TYPE "UDT_Segment"
VERSION : 0.1
   STRUCT
      MC_No_new : Byte := B#16#0;
      MC_No_old : Byte := B#16#0;
      Adresse_Peripherie : Word := W#16#0;
      Stationnumber : Byte := B#16#0;
      Spare_Byte_005 : Byte := B#16#0;
      Adr_Peripherie_analog : Word := W#16#0;
      Adr_Peripherie_SiemensFC : Word := W#16#0;
      Segment : "UDT_Station";
      Spare_Word_014 : Word := W#16#0;
      Spare_Word_016 : Word := W#16#0;
      Spare_Word_018 : Word := W#16#0;
      Input_from_segment : "UDT_Seg_input";
      Output_to_segment : "UDT_Seg_output";
      Siemens : "UDT_Siemens";
      Spare_Word_028 : Word := W#16#0;
      Spare_Word_030 : Word := W#16#0;
      Spare_Word_032 : Word := W#16#0;
      Spare_Word_034 : Word := W#16#0;
      Spare_Word_036 : Word := W#16#0;
      Spare_Word_038 : Word := W#16#0;
      Analogvalue_tool : Struct
         Input_lower_tool_1 : Word;
         Input_lower_tool_2 : Word;
         Input_upper_tool_1 : Word;
         Input_upper_tool_2 : Word;
      END_STRUCT;
      Input_from_tool : "UDT_Tool_Inputs_type_1";
      Output_to_tool : "UDT_Tool_Outputs_type_1";
      State_tool : "UDT_Mould_status";
      Spare_Word_068 : Word := W#16#0;
      Spare_Word_070 : Word := W#16#0;
      Spare_Word_072 : Word := W#16#0;
      Spare_Word_074 : Word := W#16#0;
      Spare_Word_076 : Word := W#16#0;
      Spare_Word_078 : Word := W#16#0;
      Spare_Word_080 : Word := W#16#0;
      Spare_Word_082 : Word := W#16#0;
      Spare_Word_084 : Word := W#16#0;
      Spare_Word_086 : Word := W#16#0;
      Spare_Word_088 : Word := W#16#0;
      Spare_Word_090 : Word := W#16#0;
      Spare_Word_092 : Word := W#16#0;
      Spare_Word_094 : Word := W#16#0;
      Spare_Word_096 : Word := W#16#0;
      Spare_Word_098 : Word := W#16#0;
      Segment_Bits : Struct
         WW_angewaehlt : Bool;
         Teachen_angewaehlt : Bool;
         STG_Nummer_wechselt : Bool;
         Nummer_geloescht : Bool;
         Beflammen_angewaehlt : Bool;
         Flag_TT_not_in_position : Bool;
         Reserve_100_6 : Bool;
         Reserve_100_7 : Bool;
         Reserve_101_0 : Bool;
         Reserve_101_1 : Bool;
         Reserve_101_2 : Bool;
         Reserve_101_3 : Bool;
         Reserve_101_4 : Bool;
         Reserve_101_5 : Bool;
         Reserve_101_6 : Bool;
         Reserve_101_7 : Bool;
         Reserve_Word_102 : Word;
         Reserve_Word_104 : Word;
         Reserve_Word_106 : Word;
         Reserve_Word_108 : Word;
      END_STRUCT;
      State_MC : Struct
         Movement : Struct
            RequestFromOP : "UDT_Actions";
            Request : "UDT_Actions";
            Command : "UDT_Actions";
            Valve : "UDT_Actions";
            End : "UDT_Actions";
         END_STRUCT;
         Cycle : "UDT_Cycle";
         Vacuum : "UDT_Vacuum";
         Seals : Struct
            Request_seal : Struct
               "1" : Bool;
               "2" : Bool;
               "3" : Bool;
               "4" : Bool;
               "5" : Bool;
               "6" : Bool;
               "7" : Bool;
               "8" : Bool;
               "9" : Bool;
               "10" : Bool;
               "11" : Bool;
               "12" : Bool;
               "13" : Bool;
               "14" : Bool;
               "15" : Bool;
               "16" : Bool;
               "17" : Bool;
               "18" : Bool;
               "19" : Bool;
               "20" : Bool;
               "21" : Bool;
               "22" : Bool;
               "23" : Bool;
               "24" : Bool;
               "25" : Bool;
               "26" : Bool;
               "27" : Bool;
               "28" : Bool;
               "29" : Bool;
               "30" : Bool;
               "31" : Bool;
               "32" : Bool;
            END_STRUCT;
            Seal_active : Array[0..32] of Byte;
            Flow : Struct
               Act_flow_1 : Real;
               Act_flow_2 : Real;
               Act_flow_3 : Real;
               Seal_faulty : Bool;
               Spare_12_1 : Bool;
               Spare_12_2 : Bool;
               Spare_12_3 : Bool;
               Spare_12_4 : Bool;
               Spare_12_5 : Bool;
               Spare_12_6 : Bool;
               Spare_12_7 : Bool;
               Spare_13_0 : Bool;
               Spare_13_1 : Bool;
               Spare_13_2 : Bool;
               Spare_13_3 : Bool;
               Spare_13_4 : Bool;
               Spare_13_5 : Bool;
               Spare_13_6 : Bool;
               Spare_13_7 : Bool;
            END_STRUCT;
         END_STRUCT;
         Operating_panel : Struct
            State : Struct
               Hydraulic_running : Bool := false;
               without_lockings : Bool := false;
               Spare_0_2 : Bool;
               Spare_0_3 : Bool;
               Spare_0_4 : Bool;
               Spare_0_5 : Bool;
               Spare_0_6 : Bool;
               Spare_0_7 : Bool;
               Act_step_program : Int := 0;   // Running, interupted or, for tool change: finished, running
               State_act_program : Int := 0;
               Act_operating_hours : Int := 0;
               Movement_blocked : Int := 0;
               Movement_condition_missing : Int := 0;
               Code_tool_01_actual : Int := 0;
               Code_tool_02_actual : Int := 0;
               Act_program : Int := 0;
               CounterMCCycles : DInt := L#1;
               DayCounterMCCycles : DInt := L#1;
               Act_cycle_time : Int := 0;
               Last_cycle_time : Int;
               Data_actual_MC : Int := 1;
               ProgStepNo : Int := 0;
               ProgType : Int := 5;
               Start_VNC : Bool := false;   // Bit to start the VNC viewer from PLC
               Fault_groupe_1_active : Bool := false;
               Fault_groupe_2_active : Bool := false;
               Fault_groupe_3_active : Bool := false;
               Fault_groupe_4_active : Bool := false;
               Check_USB : Bool := false;
               Spare_38_6 : Bool;
               Spare_38_7 : Bool;
            END_STRUCT;
            Set : Struct
               Insert_prog_line : Bool := false;
               Delete_prog_line : Bool := false;
               Movement_requested : Bool := false;
               Spare_0_3 : Bool := false;
               Spare_0_4 : Bool := false;
               Spare_0_5 : Bool := false;
               Request_search_missing_mov_cond : Bool := false;
               Search_missing_mov_cond : Bool := false;
               Start_loading_files : Bool := false;   // Starting loading files TP
               Loading_finished_TP : Bool := false;   // Loading finished TP (script finish)
               Loading_finished_PLC : Bool := false;   // Loading finished PLC (data in the plc)
               Request_write : Bool := false;   // Request signal to plc to write the next data block
               Release_write : Bool := false;   // Release signal to HMI (Script) to write the next data block
               Spare_1_5 : Bool := false;
               Spare_1_6 : Bool := false;
               Quit_fault : Bool := false;
               Selected_datablock : Int := 17;
               Selected_prog_line : Int := 49;
               Data_select : Int := 0;
               Data_actual : Int := 0;
               Selected_Axis : Int;
               User_level : Int;   // User level from HMI
               Spare_48_0 : Bool;
               Jog_axis_slow : Bool;   // Slow jog mode for referencing
               Jog_axis : Bool := false;
               Simmulate_tool : Bool := false;   // Simulate a tool. Reset in OB100! Only for testing
               Toggle_Lebensbit : Bool := false;
               Test_run_IBN : Bool;   // Test run for commisioning
               Spare_10_6 : Bool;
               Spare_10_7 : Bool;
               Act_file_name : String[30];
            END_STRUCT;
         END_STRUCT;
         Act_times : Struct
            Reaction_time_1 : Time;
            Reaction_time_2 : Time := T#0ms;
            Reaction_time_3 : Time := T#0ms;
            Reaction_time_4 : Time := T#0ms;
            Reaction_time_5 : Time := T#0ms;
            Reaction_time_6 : Time := T#0ms;
            Time_befor_degasing_tool_1 : Time := T#0ms;
            Degasing_time_tool_1 : Time := T#0ms;
            Time_befor_degasing_tool_2 : Time := T#0ms;
            Degasing_time_tool_2 : Time := T#0ms;
            Time_befor_degasing_tool_3 : Time := T#0ms;
            Degasing_time_tool_3 : Time := T#0ms;
            Time_befor_degasing_tool_4 : Time := T#0ms;
            Degasing_time_tool_4 : Time := T#0ms;
            Time_befor_degasing_tool_5 : Time := T#0ms;
            Degasing_time_tool_5 : Time := T#0ms;
            Time_befor_degasing_tool_6 : Time := T#0ms;
            Degasing_time_tool_6 : Time := T#0ms;
            Waiting_time_1 : Time := T#0ms;
            Waiting_time_2 : Time := T#0ms;
            Waiting_time_3 : Time := T#0ms;
            Waiting_time_4 : Time := T#0ms;
            Waiting_time_5 : Time := T#0ms;
            Waiting_time_6 : Time := T#0ms;
            Test_vacuum_circit_1 : Time := T#0ms;   // Dauer des Vakuumtestes für den Vakuumkreis 01
            Test_vacuum_circit_2 : Time := T#0ms;   // Dauer des Vakuumtestes für den Vakuumkreis 02
            Test_vacuum_circit_3 : Time := T#0ms;   // Dauer des Vakuumtestes für den Vakuumkreis 03
            Test_vacuum_circit_4 : Time := T#0ms;   // Dauer des Vakuumtestes für den Vakuumkreis 04
            Test_vacuum_circit_5 : Time := T#0ms;   // Dauer des Vakuumtestes für den Vakuumkreis 05
            Test_vacuum_circit_6 : Time := T#0ms;   // Dauer des Vakuumtestes für den Vakuumkreis 06
            Release_vacuum : Time := T#0ms;
            Switch_off_delay_vacuum_pump : Time := T#0ms;   // switch off delay for vacuum pump
            Switch_off_delay_exhaust : Time := T#0ms;   // Ausschaltverzögerung Klappe Absaugung
            Stopwatch : Time := T#0ms;
            Spare_35 : Time := T#0ms;
            Spare_36 : Time := T#0ms;
            Spare_37 : Time := T#0ms;
            Spare_38 : Time := T#0ms;
            Spare_39 : Time := T#0ms;
            Spare_40 : Time := T#0ms;
            Spare_41 : Time := T#0ms;
            Spare_42 : Time := T#0ms;
            Spare_43 : Time := T#0ms;
         END_STRUCT;
         Temperature : Struct
            Actvalue : Array[0..16] of Int;
            State : Struct
               Temp_ON : Array[0..16] of Int;
               Temp_OFF : Array[0..16] of Int;
               Heating_active_area : Array[0..16] of Bool;
            END_STRUCT;
            Faults : Struct
               F_Sensor_Temp : Array[0..16] of Bool;   // Broken wire or no sensor
               Warn_Min_Temp : Array[0..16] of Bool;   // Warning out of minimum temperature
               Tol_Min_Temp : Array[0..16] of Bool;   // Alarm out of minimum temperature
               Warn_Max_Temp : Array[0..16] of Bool;   // Warning out of maximum temperature
               Tol_Max_Temp : Array[0..16] of Bool;   // Alarm out of maximum temperature
            END_STRUCT;
            Control : Struct
               FP_heating_on_Button : Bool;
               FP_heating_off_Button : Bool;
               FP_heating_on_automatic : Bool;
               FP_heating_off_automatic : Bool;
               FP_heating_on_timecontrol : Bool;
               FP_heating_off_timecontrol : Bool;
               HF_heating_on_Button : Bool;
               HF_heating_off_Button : Bool;
               HF_heating_on_automatic : Bool;
               HF_heating_off_automatic : Bool;
               HF_heating_on_timecontrol : Bool;
               HF_heating_off_timecontrol : Bool;
               Heating_ON_Button : Bool;   // Heizungen ein über Button
               Heating_ON_timecontrol : Bool;   // Heizungen ein von Zeitschaltuhr
               Heating_ON : Bool;   // Heizungen einschalten
               Spare : Bool;
            END_STRUCT;
         END_STRUCT;
         Buttons : Struct
            OnOff : Struct
               OnOff_1 : Bool;   // Taster zum Ein/Ausschalten der Aggregate
               OnOff_2 : Bool;
               OnOff_3 : Bool;
               OnOff_4 : Bool;
               OnOff_5 : Bool;
               OnOff_6 : Bool;
               OnOff_7 : Bool;
               OnOff_8 : Bool;
               OnOff_9 : Bool;
               OnOff_10 : Bool;
               OnOff_11 : Bool;
               OnOff_12 : Bool;
               OnOff_13 : Bool;
               OnOff_14 : Bool;
               OnOff_15 : Bool;
               OnOff_16 : Bool;
               OnOff_17 : Bool;
               OnOff_18 : Bool;
               OnOff_19 : Bool;
               OnOff_20 : Bool;
               OnOff_21 : Bool;
               OnOff_22 : Bool;
               OnOff_23 : Bool;
               OnOff_24 : Bool;
               OnOff_25 : Bool;
               OnOff_26 : Bool;
               OnOff_27 : Bool;
               OnOff_28 : Bool;
               OnOff_29 : Bool;
               OnOff_30 : Bool;
               OnOff_31 : Bool;
               OnOff_32 : Bool;
            END_STRUCT;
            DisplayStatus : Array[0..31] of Byte;   // Statusbytes zur Anzeige für Schalter
         END_STRUCT;
         Tool_1 : Struct
            HF_mould_exist : Bool := true;
            Mould_exist : Bool := true;
            Only_this_mould_active : Bool := true;
            closed : Bool := false;
            Reaction_time_active_1 : Bool := false;
            Reaction_time_active_2 : Bool := false;
            Reaction_time_active_3 : Bool := false;
            Reaction_time_active_4 : Bool := false;
            Reaction_time_active_5 : Bool := false;
            Reaction_time_active_6 : Bool := false;
            Start_reaction_test : Bool := false;
            Reaction_time_started : Bool := false;
            Delete_in_out_puts : Bool := false;
            Spare_1_5 : Bool := false;
            Spare_1_6 : Bool := false;
            Reaction_time_active : Bool := false;
            Act_closing_pressure : Int := 0;
            Waiting_time_active_1 : Bool := false;
            Waiting_time_active_2 : Bool := false;
            Waiting_time_active_3 : Bool := false;
            Waiting_time_active_4 : Bool := false;
            Waiting_time_active_5 : Bool := false;
            Waiting_time_active_6 : Bool := false;
            Spare_4_6 : Bool := false;
            Spare_4_7 : Bool := false;
            foamed : Bool := false;
            flamed : Bool := false;
            Spare_5_2 : Bool := false;
            Spare_5_3 : Bool := false;
            Spare_5_4 : Bool := false;
            Spare_5_5 : Bool := false;
            Spare_5_6 : Bool := false;
            Spare_5_7 : Bool := false;
            Spare_6 : Word := 16#0000;
            Spare_8 : Word := 16#0000;
            Spare_10 : Word := 16#0000;
            Spare_12 : Word := 16#0000;
            Tool_code : "UDT_Freigabecheck";
         END_STRUCT;
         Tool_2 : Struct
            HF_mould_exist : Bool := true;
            Mould_exist : Bool := true;
            Only_this_mould_active : Bool := true;
            closed : Bool := false;
            Reaction_time_active_1 : Bool := false;
            Reaction_time_active_2 : Bool := false;
            Reaction_time_active_3 : Bool := false;
            Reaction_time_active_4 : Bool := false;
            Reaction_time_active_5 : Bool := false;
            Reaction_time_active_6 : Bool := false;
            Start_reaction_test : Bool := false;
            Reaction_time_started : Bool := false;
            Spare_1_4 : Bool := false;
            Spare_1_5 : Bool := false;
            Spare_1_6 : Bool := false;
            Reaction_time_active : Bool := false;
            Act_closing_pressure : Int := 0;
            Waiting_time_active_1 : Bool := false;
            Waiting_time_active_2 : Bool := false;
            Waiting_time_active_3 : Bool := false;
            Waiting_time_active_4 : Bool := false;
            Waiting_time_active_5 : Bool := false;
            Waiting_time_active_6 : Bool := false;
            Spare_4_6 : Bool := false;
            Spare_4_7 : Bool := false;
            foamed : Bool := false;
            flamed : Bool := false;
            Spare_5_2 : Bool := false;
            Spare_5_3 : Bool := false;
            Spare_5_4 : Bool := false;
            Spare_5_5 : Bool := false;
            Spare_5_6 : Bool := false;
            Spare_5_7 : Bool := false;
            Spare_6 : Word := 16#0000;
            Spare_8 : Word := 16#0000;
            Spare_10 : Word := 16#0000;
            Spare_12 : Word := 16#0000;
            Tool_code : "UDT_Freigabecheck";
         END_STRUCT;
         Tool_Motion : Struct
            Tool_movement_WP : Array[0..32] of "UDT_Motion";
            Tool_movement_BP : Array[0..32] of "UDT_Motion";
         END_STRUCT;
         MC_Motion : Struct
            MC_movement_WP : Array[0..32] of "UDT_Motion";
            MC_movement_BP : Array[0..32] of "UDT_Motion";
         END_STRUCT;
         IF_PU : Struct
            Bit_1 : Bool := FALSE;
            Bit_2 : Bool := FALSE;
            Bit_3 : Bool := FALSE;
            Bit_4 : Bool := FALSE;
            Bit_5 : Bool := FALSE;
            Bit_6 : Bool := FALSE;
            Bit_7 : Bool := FALSE;
            Bit_8 : Bool := FALSE;
            Bit_9 : Bool := FALSE;
            Bit_10 : Bool := FALSE;
            Bit_11 : Bool := FALSE;
            Bit_12 : Bool := FALSE;
            Bit_13 : Bool := FALSE;
            Bit_14 : Bool := FALSE;
            Bit_15 : Bool := FALSE;
            Bit_16 : Bool := FALSE;
            Word_1 : Bool := FALSE;
            Word_2 : Bool := FALSE;
         END_STRUCT;
         Toolchange : Struct
            State : Struct
               Tool_unlocked : Bool;   // --> panel for PopUp
               Tool_locked : Bool;   // --> panel for PopUp
               Profibus_disconnected : Bool;   // <- panel to carry on unlock cycle
               Water_Air_disconnected : Bool;   // <- panel to carry on unlock cycle
               Profibus_connected : Bool;   // <- panel to carry on lock cycle
               Water_Air_connected : Bool;   // <- panel to carry on lock cycle
               HF_tool_unlocked : Bool;
               HF_tool_locked : Bool;
               Semi_automatic_tool_change_active : Bool;
               Reset_light_barrier : Bool;
               Spare_1_2 : Bool;
               Spare_1_3 : Bool;
               Spare_1_4 : Bool;
               Spare_1_5 : Bool;
               Spare_1_6 : Bool;
               Spare_1_7 : Bool;
            END_STRUCT;
            Display : Struct
               Step_0 : Bool;
               Step_1 : Bool;
               Step_2 : Bool;
               Step_3 : Bool;
               Step_4 : Bool;
               Step_5 : Bool;
               Step_6 : Bool;
               Step_7 : Bool;
               Step_8 : Bool;
               Step_9 : Bool;
               Step_10 : Bool;
               Step_11 : Bool;
               Step_12 : Bool;
               Step_13 : Bool;
               Step_14 : Bool;
               Step_15 : Bool;
            END_STRUCT;
         END_STRUCT;
         "E-axis_state" : Array[0..4] of Struct
            Target_Pos_WP : Real;   // Position 1
            Target_Pos_PreWP : Real;   // Position 2
            Target_Pos_PreBP : Real;   // Position 3
            Target_Pos_BP : Real;   // Position 4
            Act_Pos : Real;
            Act_Speed : Real;
            Act_Flt : Word;   // SinaPos
            Reference_position : Bool;   // Reference sensor coverd
            HF_Reference_position : Bool;
            Request_Reference : Bool;
            Start_transfer : Bool;
            FB_was_busy : Bool;   // Helpflag that the FB was once busy
            Spare_26_5 : Bool;
            Spare_26_6 : Bool;
            Spare_26_7 : Bool;
            Profil_number : DInt;
            ErrorID : DWord;   // SinaPara
            DiagID : Word;   // SinaPara
            Error_active : Bool;
            DiagError_active : Bool;
            Spare_38_0_2 : Bool;
            Spare_38_0_3 : Bool;
            Spare_38_0_4 : Bool;
            Spare_38_0_5 : Bool;
            Spare_38_0_6 : Bool;
            Spare_38_0_7 : Bool;
            Spare_39 : Byte;
            Spare_40 : DInt;
            Spare_44 : DInt;
            Faults : Struct
               FLT_1 : Bool;   // Error code xxxx : Störung xxxxxxxxxxxxxx
               FLT_2 : Bool;   // Error code xxxx : Störung xxxxxxxxxxxxxx
               FLT_3 : Bool;   // Error code xxxx : Störung xxxxxxxxxxxxxx
               FLT_4 : Bool;   // Error code xxxx : Störung xxxxxxxxxxxxxx
               FLT_5 : Bool;   // Error code xxxx : Störung xxxxxxxxxxxxxx
               FLT_6 : Bool;   // Error code xxxx : Störung xxxxxxxxxxxxxx
               FLT_7 : Bool;   // Error code xxxx : Störung xxxxxxxxxxxxxx
               FLT_8 : Bool;   // Error code xxxx : Störung xxxxxxxxxxxxxx
               FLT_9 : Bool;   // Error code xxxx : Störung xxxxxxxxxxxxxx
               FLT_10 : Bool;   // Error code xxxx : Störung xxxxxxxxxxxxxx
               FLT_11 : Bool;   // Error code xxxx : Störung xxxxxxxxxxxxxx
               FLT_12 : Bool;   // Error code xxxx : Störung xxxxxxxxxxxxxx
               FLT_13 : Bool;   // Error code xxxx : Störung xxxxxxxxxxxxxx
               FLT_14 : Bool;   // Error code xxxx : Störung xxxxxxxxxxxxxx
               FLT_15 : Bool;   // Error code xxxx : Störung xxxxxxxxxxxxxx
               FLT_16 : Bool;   // Error code xxxx : Störung xxxxxxxxxxxxxx
               FLT_17 : Bool;   // Error code xxxx : Störung xxxxxxxxxxxxxx
               FLT_18 : Bool;   // Error code xxxx : Störung xxxxxxxxxxxxxx
               FLT_19 : Bool;   // Error code xxxx : Störung xxxxxxxxxxxxxx
               FLT_20 : Bool;   // Error code xxxx : Störung xxxxxxxxxxxxxx
               FLT_21 : Bool;   // Error code xxxx : Störung xxxxxxxxxxxxxx
               FLT_22 : Bool;   // Error code xxxx : Störung xxxxxxxxxxxxxx
               FLT_23 : Bool;   // Error code xxxx : Störung xxxxxxxxxxxxxx
               FLT_24 : Bool;   // Error code xxxx : Störung xxxxxxxxxxxxxx
            END_STRUCT;
         END_STRUCT;
         Cycle_counter : Struct
            Set : Struct
               Set_counter : Array[0..4] of DInt;
               Reset_1 : Bool;   // Stückzahl zurücksetzen
               Reset_2 : Bool;   // Stückzahl zurücksetzen
               Reset_3 : Bool;   // Stückzahl zurücksetzen
               Reset_4 : Bool;   // Stückzahl zurücksetzen
               Spare_8_4 : Bool;
               Spare_8_5 : Bool;
               Spare_8_6 : Bool;
               Spare_8_7 : Bool;
            END_STRUCT;
            State : Struct
               Act_Counter_IO : Array[0..4] of DInt;
               Act_Counter_NIO : Array[0..4] of DInt;
               Target_reached_1 : Bool;   // Stückzahl erreicht
               Target_reached_2 : Bool;   // Stückzahl erreicht
               Target_reached_3 : Bool;   // Stückzahl erreicht
               Target_reached_4 : Bool;   // Stückzahl erreicht
               Spare_8_4 : Bool;
               Spare_8_5 : Bool;
               Spare_8_6 : Bool;
               Spare_8_7 : Bool;
            END_STRUCT;
         END_STRUCT;
      END_STRUCT;
   END_STRUCT;
   // State_MC.Tool_2.Tool_code.Number_from_PU := 16#00;
   // State_MC.Tool_2.Tool_code.Spare_0_7 := false;
   // State_MC.Tool_2.Tool_code.Spare_0_6 := false;
   // State_MC.Tool_2.Tool_code.FLT_Number_in_PU_nOK := false;
   // State_MC.Tool_2.Tool_code.FLT_number_too_big := false;
   // State_MC.Tool_2.Tool_code.FLT_parity_bit := false;
   // State_MC.Tool_2.Tool_code.FLT_no_number := false;
   // State_MC.Tool_2.Tool_code.Spare_0_1 := false;
   // State_MC.Tool_2.Tool_code.HF_cycle := false;
   // State_MC.Tool_1.Tool_code.Number_from_PU := 16#00;
   // State_MC.Tool_1.Tool_code.Spare_0_7 := false;
   // State_MC.Tool_1.Tool_code.Spare_0_6 := false;
   // State_MC.Tool_1.Tool_code.FLT_Number_in_PU_nOK := false;
   // State_MC.Tool_1.Tool_code.FLT_number_too_big := false;
   // State_MC.Tool_1.Tool_code.FLT_parity_bit := false;
   // State_MC.Tool_1.Tool_code.FLT_no_number := false;
   // State_MC.Tool_1.Tool_code.Spare_0_1 := false;
   // State_MC.Tool_1.Tool_code.HF_cycle := false;
   // State_MC.Vacuum.Ready_and_okay := false;
   // State_MC.Vacuum.Motor_Dreieck := false;
   // State_MC.Vacuum.Motor_Stern := false;
   // State_MC.Vacuum.Spare_1_4 := false;
   // State_MC.Vacuum.Spare_1_3 := false;
   // State_MC.Vacuum.Spare_1_2 := false;
   // State_MC.Vacuum.Request := false;
   // State_MC.Vacuum.Flag_T_ON := false;
   // State_MC.Vacuum.Spare_0_7 := false;
   // State_MC.Vacuum.Spare_0_6 := false;
   // State_MC.Vacuum.Spare_0_5 := false;
   // State_MC.Vacuum.FLT_lock_start := false;
   // State_MC.Vacuum.FLT_filter := false;
   // State_MC.Vacuum.FLT_presure_reached := false;
   // State_MC.Vacuum.FLT_min_level_oil := false;
   // State_MC.Vacuum.FLT_motor_protection := false;
   // State_MC.Cycle.DB_Zeiger := 0;
   // State_MC.Cycle.Request_homeposition := false;
   // State_MC.Cycle.MC_in_Homeposition := false;
   // State_MC.Cycle.FP_start_Homepos_2 := false;
   // State_MC.Cycle.FP_start_Homepos_1 := false;
   // State_MC.Cycle.Homepos_active := false;
   // State_MC.Cycle.Homepos_running := false;
   // State_MC.Cycle.Cycle_lief := false;
   // State_MC.Cycle.Cycleende := false;
   // State_MC.Cycle.Spare_0_3 := false;
   // State_MC.Cycle.FP_start_Cycle := false;
   // State_MC.Cycle.Cycle_active := false;
   // State_MC.Cycle.Cycle_running := false;
   // State_MC.Movement.RequestFromOP.MCMovement01WP := FALSE;
   // State_MC.Movement.RequestFromOP.MCMovement02WP := FALSE;
   // State_MC.Movement.RequestFromOP.MCMovement03WP := FALSE;
   // State_MC.Movement.RequestFromOP.MCMovement04WP := FALSE;
   // State_MC.Movement.RequestFromOP.MCMovement05WP := FALSE;
   // State_MC.Movement.RequestFromOP.MCMovement06WP := FALSE;
   // State_MC.Movement.RequestFromOP.MCMovement07WP := FALSE;
   // State_MC.Movement.RequestFromOP.MCMovement08WP := FALSE;
   // State_MC.Movement.RequestFromOP.MCMovement09WP := FALSE;
   // State_MC.Movement.RequestFromOP.MCMovement10WP := FALSE;
   // State_MC.Movement.RequestFromOP.MCMovement11WP := FALSE;
   // State_MC.Movement.RequestFromOP.MCMovement12WP := FALSE;
   // State_MC.Movement.RequestFromOP.MCMovement13WP := FALSE;
   // State_MC.Movement.RequestFromOP.MCMovement14WP := FALSE;
   // State_MC.Movement.RequestFromOP.MCMovement15WP := FALSE;
   // State_MC.Movement.RequestFromOP.MCMovement16WP := FALSE;
   // State_MC.Movement.RequestFromOP.MCMovement17WP := FALSE;
   // State_MC.Movement.RequestFromOP.MCMovement18WP := FALSE;
   // State_MC.Movement.RequestFromOP.MCMovement19WP := FALSE;
   // State_MC.Movement.RequestFromOP.MCMovement20WP := FALSE;
   // State_MC.Movement.RequestFromOP.MCMovement21WP := FALSE;
   // State_MC.Movement.RequestFromOP.MCMovement22WP := FALSE;
   // State_MC.Movement.RequestFromOP.MCMovement23WP := FALSE;
   // State_MC.Movement.RequestFromOP.MCMovement24WP := FALSE;
   // State_MC.Movement.RequestFromOP.MCMovement25WP := FALSE;
   // State_MC.Movement.RequestFromOP.MCMovement26WP := FALSE;
   // State_MC.Movement.RequestFromOP.MCMovement27WP := FALSE;
   // State_MC.Movement.RequestFromOP.MCMovement28WP := FALSE;
   // State_MC.Movement.RequestFromOP.MCMovement29WP := FALSE;
   // State_MC.Movement.RequestFromOP.MCMovement30WP := FALSE;
   // State_MC.Movement.RequestFromOP.MCMovement31WP := FALSE;
   // State_MC.Movement.RequestFromOP.MCMovement32WP := FALSE;
   // State_MC.Movement.RequestFromOP.MCMovement01BP := FALSE;
   // State_MC.Movement.RequestFromOP.MCMovement02BP := FALSE;
   // State_MC.Movement.RequestFromOP.MCMovement03BP := FALSE;
   // State_MC.Movement.RequestFromOP.MCMovement04BP := FALSE;
   // State_MC.Movement.RequestFromOP.MCMovement05BP := FALSE;
   // State_MC.Movement.RequestFromOP.MCMovement06BP := FALSE;
   // State_MC.Movement.RequestFromOP.MCMovement07BP := FALSE;
   // State_MC.Movement.RequestFromOP.MCMovement08BP := FALSE;
   // State_MC.Movement.RequestFromOP.MCMovement09BP := FALSE;
   // State_MC.Movement.RequestFromOP.MCMovement10BP := FALSE;
   // State_MC.Movement.RequestFromOP.MCMovement11BP := FALSE;
   // State_MC.Movement.RequestFromOP.MCMovement12BP := FALSE;
   // State_MC.Movement.RequestFromOP.MCMovement13BP := FALSE;
   // State_MC.Movement.RequestFromOP.MCMovement14BP := FALSE;
   // State_MC.Movement.RequestFromOP.MCMovement15BP := FALSE;
   // State_MC.Movement.RequestFromOP.MCMovement16BP := FALSE;
   // State_MC.Movement.RequestFromOP.MCMovement17BP := FALSE;
   // State_MC.Movement.RequestFromOP.MCMovement18BP := FALSE;
   // State_MC.Movement.RequestFromOP.MCMovement19BP := FALSE;
   // State_MC.Movement.RequestFromOP.MCMovement20BP := FALSE;
   // State_MC.Movement.RequestFromOP.MCMovement21BP := FALSE;
   // State_MC.Movement.RequestFromOP.MCMovement22BP := FALSE;
   // State_MC.Movement.RequestFromOP.MCMovement23BP := FALSE;
   // State_MC.Movement.RequestFromOP.MCMovement24BP := FALSE;
   // State_MC.Movement.RequestFromOP.MCMovement25BP := FALSE;
   // State_MC.Movement.RequestFromOP.MCMovement26BP := FALSE;
   // State_MC.Movement.RequestFromOP.MCMovement27BP := FALSE;
   // State_MC.Movement.RequestFromOP.MCMovement28BP := FALSE;
   // State_MC.Movement.RequestFromOP.MCMovement29BP := FALSE;
   // State_MC.Movement.RequestFromOP.MCMovement30BP := FALSE;
   // State_MC.Movement.RequestFromOP.MCMovement31BP := FALSE;
   // State_MC.Movement.RequestFromOP.MCMovement32BP := FALSE;
   // State_MC.Movement.RequestFromOP.MouldMovement01WP := FALSE;
   // State_MC.Movement.RequestFromOP.MouldMovement02WP := FALSE;
   // State_MC.Movement.RequestFromOP.MouldMovement03WP := FALSE;
   // State_MC.Movement.RequestFromOP.MouldMovement04WP := FALSE;
   // State_MC.Movement.RequestFromOP.MouldMovement05WP := FALSE;
   // State_MC.Movement.RequestFromOP.MouldMovement06WP := FALSE;
   // State_MC.Movement.RequestFromOP.MouldMovement07WP := FALSE;
   // State_MC.Movement.RequestFromOP.MouldMovement08WP := FALSE;
   // State_MC.Movement.RequestFromOP.MouldMovement09WP := FALSE;
   // State_MC.Movement.RequestFromOP.MouldMovement10WP := FALSE;
   // State_MC.Movement.RequestFromOP.MouldMovement11WP := FALSE;
   // State_MC.Movement.RequestFromOP.MouldMovement12WP := FALSE;
   // State_MC.Movement.RequestFromOP.MouldMovement13WP := FALSE;
   // State_MC.Movement.RequestFromOP.MouldMovement14WP := FALSE;
   // State_MC.Movement.RequestFromOP.MouldMovement15WP := FALSE;
   // State_MC.Movement.RequestFromOP.MouldMovement16WP := FALSE;
   // State_MC.Movement.RequestFromOP.MouldMovement17WP := FALSE;
   // State_MC.Movement.RequestFromOP.MouldMovement18WP := FALSE;
   // State_MC.Movement.RequestFromOP.MouldMovement19WP := FALSE;
   // State_MC.Movement.RequestFromOP.MouldMovement20WP := FALSE;
   // State_MC.Movement.RequestFromOP.MouldMovement21WP := FALSE;
   // State_MC.Movement.RequestFromOP.MouldMovement22WP := FALSE;
   // State_MC.Movement.RequestFromOP.MouldMovement23WP := FALSE;
   // State_MC.Movement.RequestFromOP.MouldMovement24WP := FALSE;
   // State_MC.Movement.RequestFromOP.MouldMovement25WP := FALSE;
   // State_MC.Movement.RequestFromOP.MouldMovement26WP := FALSE;
   // State_MC.Movement.RequestFromOP.MouldMovement27WP := FALSE;
   // State_MC.Movement.RequestFromOP.MouldMovement28WP := FALSE;
   // State_MC.Movement.RequestFromOP.MouldMovement29WP := FALSE;
   // State_MC.Movement.RequestFromOP.MouldMovement30WP := FALSE;
   // State_MC.Movement.RequestFromOP.MouldMovement31WP := FALSE;
   // State_MC.Movement.RequestFromOP.MouldMovement32WP := FALSE;
   // State_MC.Movement.RequestFromOP.MouldMovement01BP := FALSE;
   // State_MC.Movement.RequestFromOP.MouldMovement02BP := FALSE;
   // State_MC.Movement.RequestFromOP.MouldMovement03BP := FALSE;
   // State_MC.Movement.RequestFromOP.MouldMovement04BP := FALSE;
   // State_MC.Movement.RequestFromOP.MouldMovement05BP := FALSE;
   // State_MC.Movement.RequestFromOP.MouldMovement06BP := FALSE;
   // State_MC.Movement.RequestFromOP.MouldMovement07BP := FALSE;
   // State_MC.Movement.RequestFromOP.MouldMovement08BP := FALSE;
   // State_MC.Movement.RequestFromOP.MouldMovement09BP := FALSE;
   // State_MC.Movement.RequestFromOP.MouldMovement10BP := FALSE;
   // State_MC.Movement.RequestFromOP.MouldMovement11BP := FALSE;
   // State_MC.Movement.RequestFromOP.MouldMovement12BP := FALSE;
   // State_MC.Movement.RequestFromOP.MouldMovement13BP := FALSE;
   // State_MC.Movement.RequestFromOP.MouldMovement14BP := FALSE;
   // State_MC.Movement.RequestFromOP.MouldMovement15BP := FALSE;
   // State_MC.Movement.RequestFromOP.MouldMovement16BP := FALSE;
   // State_MC.Movement.RequestFromOP.MouldMovement17BP := FALSE;
   // State_MC.Movement.RequestFromOP.MouldMovement18BP := FALSE;
   // State_MC.Movement.RequestFromOP.MouldMovement19BP := FALSE;
   // State_MC.Movement.RequestFromOP.MouldMovement20BP := FALSE;
   // State_MC.Movement.RequestFromOP.MouldMovement21BP := FALSE;
   // State_MC.Movement.RequestFromOP.MouldMovement22BP := FALSE;
   // State_MC.Movement.RequestFromOP.MouldMovement23BP := FALSE;
   // State_MC.Movement.RequestFromOP.MouldMovement24BP := FALSE;
   // State_MC.Movement.RequestFromOP.MouldMovement25BP := FALSE;
   // State_MC.Movement.RequestFromOP.MouldMovement26BP := FALSE;
   // State_MC.Movement.RequestFromOP.MouldMovement27BP := FALSE;
   // State_MC.Movement.RequestFromOP.MouldMovement28BP := FALSE;
   // State_MC.Movement.RequestFromOP.MouldMovement29BP := FALSE;
   // State_MC.Movement.RequestFromOP.MouldMovement30BP := FALSE;
   // State_MC.Movement.RequestFromOP.MouldMovement31BP := FALSE;
   // State_MC.Movement.RequestFromOP.MouldMovement32BP := FALSE;
   // State_MC.Movement.RequestFromOP.ShotPreparation := FALSE;
   // State_MC.Movement.RequestFromOP.ShotEnable := FALSE;
   // State_MC.Movement.RequestFromOP.ShotEnd := FALSE;
   // State_MC.Movement.RequestFromOP.StartReactionTime := FALSE;
   // State_MC.Movement.RequestFromOP.WaitReactionTime := FALSE;
   // State_MC.Movement.RequestFromOP.Spare134 := FALSE;
   // State_MC.Movement.RequestFromOP.Spare135 := FALSE;
   // State_MC.Movement.RequestFromOP.Spare136 := FALSE;
   // State_MC.Movement.RequestFromOP.Spare137 := FALSE;
   // State_MC.Movement.RequestFromOP.Spare138 := FALSE;
   // State_MC.Movement.RequestFromOP.WaitTime1 := FALSE;
   // State_MC.Movement.RequestFromOP.WaitTime2 := FALSE;
   // State_MC.Movement.RequestFromOP.WaitTime3 := FALSE;
   // State_MC.Movement.RequestFromOP.WaitTime4 := FALSE;
   // State_MC.Movement.RequestFromOP.WaitTime5 := FALSE;
   // State_MC.Movement.RequestFromOP.WaitTime6 := FALSE;
   // State_MC.Movement.RequestFromOP.StopCycle := FALSE;
   // State_MC.Movement.RequestFromOP.Spare146 := FALSE;
   // State_MC.Movement.RequestFromOP.NoFaultGroup1 := FALSE;
   // State_MC.Movement.RequestFromOP.SafetyOk := FALSE;
   // State_MC.Movement.RequestFromOP.StartWatch := FALSE;
   // State_MC.Movement.RequestFromOP.StopWatch := FALSE;
   // State_MC.Movement.RequestFromOP.Spare151 := FALSE;
   // State_MC.Movement.RequestFromOP.Spare152 := FALSE;
   // State_MC.Movement.RequestFromOP.Spare153 := FALSE;
   // // 647 more start values not shown
END_TYPE

TYPE "UDT_Station"
VERSION : 0.1
   STRUCT
      in_station_25 : Bool := FALSE;
      in_station_26 : Bool := FALSE;
      in_station_27 : Bool := FALSE;
      in_station_28 : Bool := FALSE;
      in_station_29 : Bool := FALSE;
      in_station_30 : Bool := FALSE;
      in_station_31 : Bool := FALSE;
      in_station_32 : Bool := FALSE;
      in_station_17 : Bool := FALSE;
      in_station_18 : Bool := FALSE;
      in_station_19 : Bool := FALSE;
      in_station_20 : Bool := FALSE;
      in_station_21 : Bool := FALSE;
      in_station_22 : Bool := FALSE;
      in_station_23 : Bool := FALSE;
      in_station_24 : Bool := FALSE;
      in_station_09 : Bool := FALSE;
      in_station_10 : Bool := FALSE;
      in_station_11 : Bool := FALSE;
      in_station_12 : Bool := FALSE;
      in_station_13 : Bool := FALSE;
      in_station_14 : Bool := FALSE;
      in_station_15 : Bool := FALSE;
      in_station_16 : Bool := FALSE;
      in_station_01 : Bool := FALSE;
      in_station_02 : Bool := FALSE;
      in_station_03 : Bool := FALSE;
      in_station_04 : Bool := FALSE;
      in_station_05 : Bool := FALSE;
      in_station_06 : Bool := FALSE;
      in_station_07 : Bool := FALSE;
      in_station_08 : Bool := FALSE;
   END_STRUCT;
END_TYPE

TYPE "UDT091_PouringCycleState"
TITLE = State of pouring cycle
VERSION : 0.0
   STRUCT
      Release : Bool;   // Start of shot cycle is enabled
      running : Bool;   // Shot cycle is active
      PressurizeTimeRuns : Bool;   // The time for pressure build up is running
      RmpPressurizeTimeEnd : Bool;   // Pulse time for pressure build up is finished
      PressurizeTimeFinished : Bool;   // Time for pressure build up was finished correctly -> 1 until end of cycle
      StandByTimeRuns : Bool;   // Time after shot while next start shot is possible
      RmpStandByTimeEnd : Bool;   // Pulse stand by time is finished (means that cycle is finished)
      CtrlChangeTimeRuns : Bool;   // Time for change of controller values (flow, pressure,...) runs
      RmpCtrlChangeTimeEnd : Bool;   // Pulse time for change of controller values finished
      Shotrelease : Bool;   // foaming cycle is ready for foaming (times are finished)
      ShotRuns : Bool;   // Mixinghead is open (or service shot runs)
      PulsShotend : Bool;   // Pulse shot was finished
      MHWasOpen : Bool;   // Information MH was opened
      PulseCycleEnd : Bool;   // Pulse shot cycle is finished
      SelectHydForShot : Bool;   // Request HD-valve of hydraulics
      NoReleaseDuringShot : Bool;   // shot was finished too early, because release was set to zero
      FLT_KLZ_0 : Bool;   // Fault recirculition time 0
      FLT_MaxWaittime : Bool;   // fault no shot started after maximum waiting time
      FLT_MaxShottime : Bool;   // Fault shottime too long
      FLT_OPMode : Bool;   // OP mode changed between service and shot with foaming during shot
      LastShotinTool : Bool;   // After this shot the foamingcycle of this tool (mould) is finished
      LastShotinToolFinished : Bool;
      Pulse_ToolFinished : Bool;   // Pulse last shot of tool finished
      LastStanbyTimeTool : Bool;   // Tool finished
      Stepnumber : Byte;   // Stepcounter for sequence of shot cycle
   END_STRUCT;
END_TYPE

TYPE "UDT_Seg_output"
VERSION : 0.1
   STRUCT
      O_bold_PS_lock : Bool;   // Lock parallelstroke (UMP/LMP)
      O_bold_PS_unlock : Bool;   // Unock parallelstroke (UMP/LMP)
      O_safetybold_PS_unlock : Bool;   // Unlock safety bold parallel stroke
      O_release_break_PS : Bool;   // Release break parallel stroke
      O_safetybold_UMP_unlock : Bool;   // safety bold upper mold plate unlocked
      O_Aircushion_up : Bool;   // aircushion up
      O_Aircushion_down : Bool;   // aircushion down
      O_spare_2x0_7 : Bool;
      O_MldLckLP_lock : Bool;   // Lock tool change lower plate
      O_MldLckLP_unlock : Bool;   // Unlock tool change lower plate
      O_MldLckUP_lock : Bool;   // Lock tool change upper plate
      O_MldLckUP_unlock : Bool;   // Unlock tool change upper plate
      O_MldLckUP_break : Bool;   // Release break tool change upper plate
      O_spare_2x5_5 : Bool;
      O_spare_2x5_6 : Bool;
      O_spare_2x5_7 : Bool;
   END_STRUCT;
END_TYPE

TYPE "UDT_Cycle"
VERSION : 0.0
   STRUCT
      Cycle_running : Bool;   // Poduction cycle running
      Cycle_active : Bool;   // Production cycle running and active (not interrupted)
      FP_start_Cycle : Bool;
      Spare_0_3 : Bool;
      Cycleende : Bool;
      Cycle_lief : Bool;
      Spare_0_6 : Bool;
      Request_cycle : Bool;
      Homepos_running : Bool;   // Homepos cycle running
      Homepos_active : Bool;   // Homepos cycle running and active (not interrupted)
      FP_start_Homepos_1 : Bool;
      FP_start_Homepos_2 : Bool;
      MC_in_Homeposition : Bool;
      Flag_start_home_1 : Bool;
      Flag_start_home_2 : Bool;
      Request_homeposition : Bool;
      Breakpos_running : Bool;   // Breakpos cycle running
      Breakpos_active : Bool;   // Breakpos cycle running and active (not interrupted)
      FP_start_Breakpos : Bool;
      Spare_2_3 : Bool;
      MC_in_Breakposition : Bool;
      Spare_2_5 : Bool;
      Spare_2_6 : Bool;
      Request_breakposition : Bool;
      Testshot_running : Bool;   // Testshot cycle running
      Testshot_active : Bool;   // Testshot cycle running and active (not interrupted)
      FP_start_Testshot : Bool;
      Spare_3_3 : Bool;
      MC_in_Testshotposition : Bool;
      Spare_3_5 : Bool;
      Spare_3_6 : Bool;
      Request_testshotposition : Bool;
      Flag_degassing_inflate : Bool := false;
      Flag_degassing_deflate : Bool := false;
      Flag_degassing_duration : Bool := false;
      Flag_degassing : Bool := false;
      Request_degassing : Bool := false;
      MC_was_in_degassing_position : Bool := false;
      Cycle_release : Bool := false;   // Cycle release, all condidtions are okay
      Temperature_okay : Bool := false;   // No Tolerance alarm for start cycle
      Lock_seals : Bool;   // Lock seals
      Cycle_running_TP : Bool;
      Fault_MC : Bool;
      Turn_lock : Bool;
      No_foaming : Bool;
      Delete_cycle : Bool;
      Release_production : Bool;
      Access_release_MC : Bool;
      FT_gesperrt : Bool;
      FT_angewaehlt : Bool;
      FT_Schaeumvorbereitung : Bool;
      FT_Schaeumfreigabe : Bool;
      FT_Schaeumende : Bool;
      FT_Schaeumstoerung : Bool;
      Zyklus_abbrechen : Bool;
      FT_hat_Zyklus_gestartet : Bool;
      FHM_Start_schaeumen : Bool;
      FHM_Stop_schaeumen : Bool;
      Spare_4 : Bool;
      Spare_5 : Bool;
      Spare_6 : Bool;
      Spare_7 : Bool;
      Spare_8 : Bool;
      Spare_9 : Bool;
      Spare_10 : Bool;
      Spare_11 : Bool;
      Spare_12 : Bool;
      Spare_13 : Bool;
      Spare_14 : Bool;
      Spare_15 : Bool;
      Spare_16 : Bool;
      Spare_17 : Bool;
      Spare_18 : Byte;
      DB_Zeiger : Int;
   END_STRUCT;
END_TYPE

TYPE "UDT_Motion"
VERSION : 0.0
   STRUCT
      Action_1 : Bool;
      Action_2 : Bool;
      Action_3 : Bool;
      Action_4 : Bool;
      Action_5 : Bool;
      Action_6 : Bool;
      Action_7 : Bool;
      Action_8 : Bool;
      Action_9 : Bool;
      Action_10 : Bool;
      Action_11 : Bool;
      Action_12 : Bool;
      Action_13 : Bool;
      Action_14 : Bool;
      Core_in_endposition : Bool;   // For WinCap, Jaeckl and IP (FB18)
      Opposite_position_reached : Bool;
      FLT_running_time : Bool;
      FLT_Sensor : Bool;
      FLT_Spare_2_2 : Bool;
      FLT_Spare_2_3 : Bool;
      FLT_Spare_2_4 : Bool;
      FLT_Spare_2_5 : Bool;
      FLT_Spare_2_6 : Bool;
      FLT_Spare_2_7 : Bool;
   END_STRUCT;
END_TYPE

TYPE "UDT095_MouldPressureCont"
VERSION : 0.1
   STRUCT
      FLT_UpperLimitFlow : Bool;
      FLT_LowerLimitFlow : Bool;
      FLT_Spare02 : Bool;
      FLT_Spare03 : Bool;
      FLT_Spare04 : Bool;
      FLT_Spare05 : Bool;
      Spare06 : Bool;
      Spare07 : Bool;
      WorkCycle_Flag1 : Bool;
      WorkCycle_Flag2 : Bool;
      Enableclosedloop : Bool;   // PLC-release to control the component flow at modul
      DecrementFlow : Bool;
      IncrementFlow : Bool;
      EnableFlowControl : Bool;
      Switch_Drive_ON_OFF : Bool;
      FirstSensorControlActive : Bool;
      State_Drive : Int;   // 1->Drive ON; 2->Fault Drive; 3->Drive requested but not on
      PSetValueReachedS01 : Bool;
      PSetValueReachedS02 : Bool;
      PSetValueReachedS03 : Bool;
      PSetValueReachedS04 : Bool;
      PSetValueReachedS05 : Bool;
      PSetValueReachedS06 : Bool;
      PSetValueReachedS07 : Bool;
      PSetValueReachedS08 : Bool;
      WorkFinishedS01 : Bool;
      WorkFinishedS02 : Bool;
      WorkFinishedS03 : Bool;
      WorkFinishedS04 : Bool;
      WorkFinishedS05 : Bool;
      WorkFinishedS06 : Bool;
      WorkFinishedS07 : Bool;
      WorkFinishedS08 : Bool;
      SensorActive01 : Bool;
      SensorActive02 : Bool;
      SensorActive03 : Bool;
      SensorActive04 : Bool;
      SensorActive05 : Bool;
      SensorActive06 : Bool;
      SensorActive07 : Bool;
      SensorActive08 : Bool;
   END_STRUCT;
END_TYPE

TYPE "UDT_Siemens"
AUTHOR : KT242
VERSION : 0.1
   STRUCT
      Supply_unit : Struct
         HW_ID : Hw_Any;
         Input : Struct
            "1" : Bool;
            Führung_gefordert : Bool;
            "3" : Bool;
            Vorladung_beendet : Bool;
            Netzschütz_geschlossen : Bool;
            "6" : Bool;
            "7" : Bool;
            "8" : Bool;
            Einschaltbereit : Bool;
            Betriebsbereit : Bool;
            Betrieb_freigegeben : Bool;
            Störung_wirksam : Bool;
            Kein_AUS_2_aktiv : Bool;
            "14" : Bool;
            Einschaltsperre : Bool;
            Warnung_wirksam : Bool;
         END_STRUCT;
         Output : Struct
            "1" : Bool;
            "2" : Bool;
            Führung_durch_PLC : Bool;
            "4" : Bool;
            "5" : Bool;
            "6" : Bool;
            "7" : Bool;
            "8" : Bool;
            ON : Bool;
            Kein_austrudeln : Bool;
            "11" : Bool;
            Betrieb_freigegeben : Bool;
            "13" : Bool;
            "14" : Bool;
            Einspeisung_generatorischen_Betrieb_sperren : Bool;
            Störung_quittieren : Bool;
         END_STRUCT;
      END_STRUCT;
      FC_1 : "UDT_Siemens_FC";
      FC_2 : "UDT_Siemens_FC";
      FC_3 : "UDT_Siemens_FC";
      FC_4 : "UDT_Siemens_FC";
   END_STRUCT;
END_TYPE

TYPE "UDT_Freigabecheck"
VERSION : 0.1
   STRUCT
      HF_cycle : Bool;
      Spare_0_1 : Bool;
      FLT_no_number : Bool;
      FLT_parity_bit : Bool;
      FLT_number_too_big : Bool;
      FLT_Number_in_PU_nOK : Bool;
      Spare_0_6 : Bool;
      Spare_0_7 : Bool;
      Number_from_PU : Byte;
   END_STRUCT;
END_TYPE

TYPE "UDT_MVM_Settings"
AUTHOR : KT242
VERSION : 0.1
   STRUCT
      Position : Array[1..4] of Struct
         Target : Real;   // Targetposition
         Switch_over_offset_start : Real;   // Offset from targetposition to switch to last profil
         Switch_over_offset_end : Real;   // Offset from start position with first profil
         Speed_manual : Int;   // Speed in manual mode
         Speed_automatic : Int;   // Speed in automatic mode profil 1
         Acceleration : Int;   // Acceleration profil 1
         Deceleration : Int;   // Deceleration profil 1
         Speed_automatic_2 : Int;   // Speed in automatic mode profil 2
         Acceleration_2 : Int;   // Acceleration profil 2
         Deceleration_2 : Int;   // Deceleration profil 2
         Speed_automatic_3 : Int;   // Speed in automatic mode profil 3
         Acceleration_3 : Int;   // Acceleration profil 3
         Deceleration_3 : Int;   // Deceleration profil 3
      END_STRUCT;
   END_STRUCT;
END_TYPE

TYPE "UDT2000_KM_FRA"
VERSION : 0.1
   STRUCT
      Flanke_Strobe : Bool;
      Flanke_Strobe_inv : Bool;
      Flanke_MK_Open : Bool;
      Fehler_FA_nicht_bereit : Bool;
      Fehler_keine_Nummer : Bool;   // Strobe gesetzt aber keine Nummer liegt an
      Fehler_invers : Bool;   // Die invertierte Nummer war falsch
      Fehler_PBit : Bool;   // Parity bit kam falsch
      Prg_ok : Bool;
      Start_an_PU : Bool;
      MK_open_an_PU : Bool;
      RK_vor_an_PU : Bool;
      Flanke_Res_MK_open : Bool;
      Flanke_TSE : Bool;   // Flanke für Teilschussende
      MK_war_auf : Bool;
      Imp_MK_open : Bool;
      Role_bit : Bool;
      PrgNr_Speicher : Byte;
      PrgNr_invers_Speicher : Byte;
      PrgNr_an_PU : Byte;
      "Step" : Byte;
   END_STRUCT;
END_TYPE

TYPE "UDT2001_Input_Faurecia"
VERSION : 0.1
   STRUCT
      comandstatus : Struct
         STROBE : Bool;   // 1 = Start foamcycle, foam values are valid
         STARTSHOT : Bool;   // 1 = release mixhead open
         STOP : Bool;   // 0 = stop foaming, shot abort
         CPFORWARD : Bool := FALSE;   // 1 = move cleaning piston forward (outside a foamcycle)
         Reset_Fault : Bool := FALSE;   // 1 = Acknowledge alarms
         Service : Bool := FALSE;   // 1 = Service mode selection
         RedCirc : Bool := FALSE;   // 1 = Start/ Stop reduced circulation
         Watchdog : Bool := FALSE;   // 1 = Line PLC watchdog
         Reserve6 : Byte := B#16#0;
      END_STRUCT;
      foaming_values : Struct
         shottime : DWord := DW#16#0;   // setvalue shottime in ms
         flow_C1 : Word := W#16#0;   // setvalue flow C1 in 1/10g/s
         flow_C2 : Word := W#16#0;   // setvalue flow C2 in 1/10g/s
         pressure_C1 : Word := W#16#0;   // setvalue pressure C1 in bar
         pressure_C2 : Word := W#16#0;   // setvalue pressure C2 in bar
         Reserve0 : Bool := FALSE;
         CP_AFTER_SHOT : Bool := FALSE;   // 1 = cleaning piston should move immediate after shot
         Reserve1 : Bool := FALSE;
         Reserve2 : Bool := FALSE;
         Reserve3 : Bool := FALSE;
         Reserve4 : Bool := FALSE;
         Reserve5 : Bool := FALSE;
         Reserve6 : Bool := FALSE;
         Reserve7 : Byte := B#16#0;
      END_STRUCT;
      Reserve : Struct
         Reserve1 : Word := W#16#0;
         Reserve2 : Word := W#16#0;
         Reserve3 : Word := W#16#0;
         Reserve4 : Word := W#16#0;
      END_STRUCT;
   END_STRUCT;
END_TYPE

TYPE "UDT710_Agitator"
TITLE = State of auxiliary drive